// TIA Portal project "HEAT-1-CADIZ-V30" (V20) (continued)
VAR_GLOBAL   // PLC tag table "Robot Position"
   "tcpPosIniX_00" AT %I632.0 : Bool;   // $OUT[257]
   "tcpPosIniX_01" AT %I632.1 : Bool;
   "tcpPosIniX_02" AT %I632.2 : Bool;
   "tcpPosIniX_03" AT %I632.3 : Bool;
   "tcpPosIniX_04" AT %I632.4 : Bool;
   "tcpPosIniX_05" AT %I632.5 : Bool;
   "tcpPosIniX_06" AT %I632.6 : Bool;
   "tcpPosIniX_07" AT %I632.7 : Bool;
   "tcpPosIniX_08" AT %I633.0 : Bool;
   "tcpPosIniX_09" AT %I633.1 : Bool;
   "tcpPosIniX_10" AT %I633.2 : Bool;
   "tcpPosIniX_11" AT %I633.3 : Bool;
   "tcpPosIniX_12" AT %I633.4 : Bool;
   "tcpPosIniX_13" AT %I633.5 : Bool;
   "tcpPosIniX_14" AT %I633.6 : Bool;
   "tcpPosIniX_15" AT %I633.7 : Bool;
   "tcpPosIniX_16" AT %I634.0 : Bool;
   "tcpPosIniX_17" AT %I634.1 : Bool;
   "tcpPosIniX_18" AT %I634.2 : Bool;
   "tcpPosIniX_19" AT %I634.3 : Bool;
   "tcpPosIniX_20" AT %I634.4 : Bool;
   "tcpPosIniX_21" AT %I634.5 : Bool;
   "tcpPosIniX_22" AT %I634.6 : Bool;
   "tcpPosIniX_23" AT %I634.7 : Bool;
   "tcpPosIniX_24" AT %I635.0 : Bool;
   "tcpPosIniX_25" AT %I635.1 : Bool;
   "tcpPosIniX_26" AT %I635.2 : Bool;
   "tcpPosIniX_27" AT %I635.3 : Bool;
   "tcpPosIniX_28" AT %I635.4 : Bool;
   "tcpPosIniX_29" AT %I635.5 : Bool;
   "tcpPosIniX_30" AT %I635.6 : Bool;
   "tcpPosIniX_31" AT %I635.7 : Bool;
   "tcpPosIniY_00" AT %I636.0 : Bool;
   "tcpPosIniY_01" AT %I636.1 : Bool;
   "tcpPosIniY_02" AT %I636.2 : Bool;
   "tcpPosIniY_03" AT %I636.3 : Bool;
   "tcpPosIniY_04" AT %I636.4 : Bool;
   "tcpPosIniY_05" AT %I636.5 : Bool;
   "tcpPosIniY_06" AT %I636.6 : Bool;
   "tcpPosIniY_07" AT %I636.7 : Bool;
   "tcpPosIniY_08" AT %I637.0 : Bool;
   "tcpPosIniY_09" AT %I637.1 : Bool;
   "tcpPosIniY_10" AT %I637.2 : Bool;
   "tcpPosIniY_11" AT %I637.3 : Bool;
   "tcpPosIniY_12" AT %I637.4 : Bool;
   "tcpPosIniY_13" AT %I637.5 : Bool;
   "tcpPosIniY_14" AT %I637.6 : Bool;
   "tcpPosIniY_15" AT %I637.7 : Bool;
   "tcpPosIniY_16" AT %I638.0 : Bool;
   "tcpPosIniY_17" AT %I638.1 : Bool;
   "tcpPosIniY_18" AT %I638.2 : Bool;
   "tcpPosIniY_19" AT %I638.3 : Bool;
   "tcpPosIniY_20" AT %I638.4 : Bool;
   "tcpPosIniY_21" AT %I638.5 : Bool;
   "tcpPosIniY_22" AT %I638.6 : Bool;
   "tcpPosIniY_23" AT %I638.7 : Bool;
   "tcpPosIniY_24" AT %I639.0 : Bool;
   "tcpPosIniY_25" AT %I639.1 : Bool;
   "tcpPosIniY_26" AT %I639.2 : Bool;
   "tcpPosIniY_27" AT %I639.3 : Bool;
   "tcpPosIniY_28" AT %I639.4 : Bool;
   "tcpPosIniY_29" AT %I639.5 : Bool;
   "tcpPosIniY_30" AT %I639.6 : Bool;
   "tcpPosIniY_31" AT %I639.7 : Bool;
   "tcpPosIniZ_00" AT %I640.0 : Bool;
   "tcpPosIniZ_01" AT %I640.1 : Bool;
   "tcpPosIniZ_02" AT %I640.2 : Bool;
   "tcpPosIniZ_03" AT %I640.3 : Bool;
   "tcpPosIniZ_04" AT %I640.4 : Bool;
   "tcpPosIniZ_05" AT %I640.5 : Bool;
   "tcpPosIniZ_06" AT %I640.6 : Bool;
   "tcpPosIniZ_07" AT %I640.7 : Bool;
   "tcpPosIniZ_08" AT %I641.0 : Bool;
   "tcpPosIniZ_09" AT %I641.1 : Bool;
   "tcpPosIniZ_10" AT %I641.2 : Bool;
   "tcpPosIniZ_11" AT %I641.3 : Bool;
   "tcpPosIniZ_12" AT %I641.4 : Bool;
   "tcpPosIniZ_13" AT %I641.5 : Bool;
   "tcpPosIniZ_14" AT %I641.6 : Bool;
   "tcpPosIniZ_15" AT %I641.7 : Bool;
   "tcpPosIniZ_16" AT %I642.0 : Bool;
   "tcpPosIniZ_17" AT %I642.1 : Bool;
   "tcpPosIniZ_18" AT %I642.2 : Bool;
   "tcpPosIniZ_19" AT %I642.3 : Bool;
   "tcpPosIniZ_20" AT %I642.4 : Bool;
   "tcpPosIniZ_21" AT %I642.5 : Bool;
   "tcpPosIniZ_22" AT %I642.6 : Bool;
   "tcpPosIniZ_23" AT %I642.7 : Bool;
   "tcpPosIniZ_24" AT %I643.0 : Bool;
   "tcpPosIniZ_25" AT %I643.1 : Bool;
   "tcpPosIniZ_26" AT %I643.2 : Bool;
   "tcpPosIniZ_27" AT %I643.3 : Bool;
   "tcpPosIniZ_28" AT %I643.4 : Bool;
   "tcpPosIniZ_29" AT %I643.5 : Bool;
   "tcpPosIniZ_30" AT %I643.6 : Bool;
   "tcpPosIniZ_31" AT %I643.7 : Bool;
   "e1PosIni_00" AT %I644.0 : Bool;
   "e1PosIni_01" AT %I644.1 : Bool;
   "e1PosIni_02" AT %I644.2 : Bool;
   "e1PosIni_03" AT %I644.3 : Bool;
   "e1PosIni_04" AT %I644.4 : Bool;
   "e1PosIni_05" AT %I644.5 : Bool;
   "e1PosIni_06" AT %I644.6 : Bool;
   "e1PosIni_07" AT %I644.7 : Bool;
   "e1PosIni_08" AT %I645.0 : Bool;
   "e1PosIni_09" AT %I645.1 : Bool;
   "e1PosIni_10" AT %I645.2 : Bool;
   "e1PosIni_11" AT %I645.3 : Bool;
   "e1PosIni_12" AT %I645.4 : Bool;
   "e1PosIni_13" AT %I645.5 : Bool;
   "e1PosIni_14" AT %I645.6 : Bool;
   "e1PosIni_15" AT %I645.7 : Bool;
   "e1PosIni_16" AT %I646.0 : Bool;
   "e1PosIni_17" AT %I646.1 : Bool;
   "e1PosIni_18" AT %I646.2 : Bool;
   "e1PosIni_19" AT %I646.3 : Bool;
   "e1PosIni_20" AT %I646.4 : Bool;
   "e1PosIni_21" AT %I646.5 : Bool;
   "e1PosIni_22" AT %I646.6 : Bool;
   "e1PosIni_23" AT %I646.7 : Bool;
   "e1PosIni_24" AT %I647.0 : Bool;
   "e1PosIni_25" AT %I647.1 : Bool;
   "e1PosIni_26" AT %I647.2 : Bool;
   "e1PosIni_27" AT %I647.3 : Bool;
   "e1PosIni_28" AT %I647.4 : Bool;
   "e1PosIni_29" AT %I647.5 : Bool;
   "e1PosIni_30" AT %I647.6 : Bool;
   "e1PosIni_31" AT %I647.7 : Bool;
   "tcpPosFinX_00" AT %I648.0 : Bool;
   "tcpPosFinX_01" AT %I648.1 : Bool;
   "tcpPosFinX_02" AT %I648.2 : Bool;
   "tcpPosFinX_03" AT %I648.3 : Bool;
   "tcpPosFinX_04" AT %I648.4 : Bool;
   "tcpPosFinX_05" AT %I648.5 : Bool;
   "tcpPosFinX_06" AT %I648.6 : Bool;
   "tcpPosFinX_07" AT %I648.7 : Bool;
   "tcpPosFinX_08" AT %I649.0 : Bool;
   "tcpPosFinX_09" AT %I649.1 : Bool;
   "tcpPosFinX_10" AT %I649.2 : Bool;
   "tcpPosFinX_11" AT %I649.3 : Bool;
   "tcpPosFinX_12" AT %I649.4 : Bool;
   "tcpPosFinX_13" AT %I649.5 : Bool;
   "tcpPosFinX_14" AT %I649.6 : Bool;
   "tcpPosFinX_15" AT %I649.7 : Bool;
   "tcpPosFinX_16" AT %I650.0 : Bool;
   "tcpPosFinX_17" AT %I650.1 : Bool;
   "tcpPosFinX_18" AT %I650.2 : Bool;
   "tcpPosFinX_19" AT %I650.3 : Bool;
   "tcpPosFinX_20" AT %I650.4 : Bool;
   "tcpPosFinX_21" AT %I650.5 : Bool;
   "tcpPosFinX_22" AT %I650.6 : Bool;
   "tcpPosFinX_23" AT %I650.7 : Bool;
   "tcpPosFinX_24" AT %I651.0 : Bool;
   "tcpPosFinX_25" AT %I651.1 : Bool;
   "tcpPosFinX_26" AT %I651.2 : Bool;
   "tcpPosFinX_27" AT %I651.3 : Bool;
   "tcpPosFinX_28" AT %I651.4 : Bool;
   "tcpPosFinX_29" AT %I651.5 : Bool;
   "tcpPosFinX_30" AT %I651.6 : Bool;
   "tcpPosFinX_31" AT %I651.7 : Bool;
   "tcpPosFinY_00" AT %I652.0 : Bool;
   "tcpPosFinY_01" AT %I652.1 : Bool;
   "tcpPosFinY_02" AT %I652.2 : Bool;
   "tcpPosFinY_03" AT %I652.3 : Bool;
   "tcpPosFinY_04" AT %I652.4 : Bool;
   "tcpPosFinY_05" AT %I652.5 : Bool;
   "tcpPosFinY_06" AT %I652.6 : Bool;
   "tcpPosFinY_07" AT %I652.7 : Bool;
   "tcpPosFinY_08" AT %I653.0 : Bool;
   "tcpPosFinY_09" AT %I653.1 : Bool;
   "tcpPosFinY_10" AT %I653.2 : Bool;
   "tcpPosFinY_11" AT %I653.3 : Bool;
   "tcpPosFinY_12" AT %I653.4 : Bool;
   "tcpPosFinY_13" AT %I653.5 : Bool;
   "tcpPosFinY_14" AT %I653.6 : Bool;
   "tcpPosFinY_15" AT %I653.7 : Bool;
   "tcpPosFinY_16" AT %I654.0 : Bool;
   "tcpPosFinY_17" AT %I654.1 : Bool;
   "tcpPosFinY_18" AT %I654.2 : Bool;
   "tcpPosFinY_19" AT %I654.3 : Bool;
   "tcpPosFinY_20" AT %I654.4 : Bool;
   "tcpPosFinY_21" AT %I654.5 : Bool;
   "tcpPosFinY_22" AT %I654.6 : Bool;
   "tcpPosFinY_23" AT %I654.7 : Bool;
   "tcpPosFinY_24" AT %I655.0 : Bool;
   "tcpPosFinY_25" AT %I655.1 : Bool;
   "tcpPosFinY_26" AT %I655.2 : Bool;
   "tcpPosFinY_27" AT %I655.3 : Bool;
   "tcpPosFinY_28" AT %I655.4 : Bool;
   "tcpPosFinY_29" AT %I655.5 : Bool;
   "tcpPosFinY_30" AT %I655.6 : Bool;
   "tcpPosFinY_31" AT %I655.7 : Bool;
   "tcpPosE1_01" AT %I628.0 : Bool;
   "tcpPosE1_02" AT %I628.1 : Bool;
   "tcpPosE1_03" AT %I628.2 : Bool;
   "tcpPosE1_04" AT %I628.3 : Bool;
   "tcpPosE1_05" AT %I628.4 : Bool;
   "tcpPosE1_06" AT %I628.5 : Bool;
   "tcpPosE1_07" AT %I628.6 : Bool;
   "tcpPosE1_08" AT %I628.7 : Bool;
   "tcpPosE1_09" AT %I629.0 : Bool;
   "tcpPosE1_10" AT %I629.1 : Bool;
   "tcpPosE1_11" AT %I629.2 : Bool;
   "tcpPosE1_12" AT %I629.3 : Bool;
   "tcpPosE1_13" AT %I629.4 : Bool;
   "tcpPosE1_14" AT %I629.5 : Bool;
   "tcpPosE1_15" AT %I629.6 : Bool;
   "tcpPosE1_16" AT %I629.7 : Bool;
   "tcpPosE1_17" AT %I630.0 : Bool;
   "tcpPosE1_18" AT %I630.1 : Bool;
   "tcpPosE1_19" AT %I630.2 : Bool;
   "tcpPosE1_20" AT %I630.3 : Bool;
   "tcpPosE1_21" AT %I630.4 : Bool;
   "tcpPosE1_22" AT %I630.5 : Bool;
   "tcpPosE1_23" AT %I630.6 : Bool;
   "tcpPosE1_24" AT %I630.7 : Bool;
   "tcpPosE1_25" AT %I631.0 : Bool;
   "tcpPosE1_26" AT %I631.1 : Bool;
   "tcpPosE1_27" AT %I631.2 : Bool;
   "tcpPosE1_28" AT %I631.3 : Bool;
   "tcpPosE1_29" AT %I631.4 : Bool;
   "tcpPosE1_30" AT %I631.5 : Bool;
   "tcpPosE1_31" AT %I631.6 : Bool;
   "tcpPosE1_32" AT %I631.7 : Bool;
   "tcpPosIniX_rawLe32" AT %ID632 : DWord;
   "tcpPosIniY_rawLe32" AT %ID636 : DWord;
   "tcpPosIniZ_rawLe32" AT %ID640 : DWord;
   "tcpPosFinX_rawLe32" AT %ID648 : DWord;
   "tcpPosFinY_rawLe32" AT %ID652 : DWord;
   "e1_rawLe32" AT %ID628 : DWord;
   "e1PosIni_rawLe32" AT %ID644 : DWord;
   "tcpPosFinZ_rawLe32" AT %ID656 : DWord;
   "e1PosFin_rawLe32" AT %ID660 : DWord;
END_VAR

VAR_GLOBAL   // PLC tag table "Tool Change"
   "dockSensorToolYugoInPosition" AT %I150.0 : Bool;   // DETECTOR_YUGO_LP
   "dockSensorCoverYugoClosed" AT %I150.1 : Bool;   // TAPA_CERRADA_YUGO_LP
   "dockSensorCoverOpenYugo" AT %I160.0 : Bool;   // TAPA_ABIERTA_YUGO_LP
   "dockValveV2UnlockOnYugo" AT %Q171.2 : Bool;   // SOLTAR_HERRAMIENTA_YUGO_LP / CAMBIA A FALSE
   "dockValveCoverOpenOnYugo" AT %Q170.0 : Bool;   // ABRIR_TAPA_YUGO_LP
   "dockValveCoverCloseOnYugo" AT %Q170.1 : Bool;   // CERRAR_TAPA_YUGO_LP
   "robotSensorMpsUnlocked" AT %I200.0 : Bool;   // INTERCAMBIO_DESBLOQUEADO_LR
   "robotSensorMpsLocked" AT %I200.1 : Bool;   // INTERCAMBIO_BLOQUEADO_LR
   "robotSensorMpsCoupled" AT %I200.2 : Bool;   // HERRAMIENTA_PUESTA_LR /AL COLOCAR METAL
   "robotSensorMpsCtrlAirPressureOk" AT %I200.3 : Bool;   // PRESION_CORRECTA_LR
   "toolReqId_01" AT %Q618.1 : Bool;   // INKUKA_DETECTOR_HERRAMIENTA
   "toolReqId_02" AT %Q618.2 : Bool;   // INKUKA_TAPA_CERRADA_YUGO
   "toolReqId_03" AT %Q618.3 : Bool;   // INKUKA_TAPA_ABIERTA_YUGO
   "toolReqId_04" AT %Q618.4 : Bool;   // INKUKA_INTERCAMBIO_DESBLOQUEADO
   "toolReqId_05" AT %Q618.5 : Bool;   // INKUKA_INTERCAMBIO_BLOQUEADO
   "toolReqId_06" AT %Q618.6 : Bool;   // INKUKA_HERRAMIENTA_PUESTA /AL COLOCAR util met
   "toolReqId_07" AT %Q618.7 : Bool;
   "kukaCmdUnlockMpsYugo" AT %I696.0 : Bool;   // OUTKUKA_SOLTAR_HERRAMIENTA_YUGO
   "kukaCmdOpenCover" AT %I696.1 : Bool;   // OUTKUKA_ABRIR_TAPA_YUGO
   "kukaCmdCloseCover" AT %I696.2 : Bool;   // OUTKUKA_CERRAR_TAPA_YUGO
   "V1_B14_S2" AT %Q0.0 : Bool;   // Anticolision - OPR
   "V1_B12_S4" AT %Q0.1 : Bool;   // Mps Bloqueo SIL 2
   "V2_B14_S2" AT %Q0.2 : Bool;
   "V2_B12_S4" AT %Q0.3 : Bool;
   "toolReqId_00" AT %Q618.0 : Bool;
   "toolReqId_08" AT %Q619.0 : Bool;
   "toolReqId_09" AT %Q619.1 : Bool;
   "toolReqId_10" AT %Q619.2 : Bool;
   "toolReqId_11" AT %Q619.3 : Bool;
   "toolReqId_12" AT %Q619.4 : Bool;
   "toolReqId_13" AT %Q619.5 : Bool;
   "toolReqId_14" AT %Q619.6 : Bool;
   "toolReqId_15" AT %Q619.7 : Bool;
   "toolReqId" AT %QW618 : Word;
   "baseReqId" AT %QW620 : Word;
   "kukaFeedbackDockToolYugoInPosition" AT %Q696.4 : Bool;   // $IN[773]
   "kukaFeedbackDockYugoCoverClosed" AT %Q696.5 : Bool;
   "kukaFeedbackDockYugoCoverOpen" AT %Q696.6 : Bool;
   "kukaFeedbackRobotMpsUnlocked" AT %Q696.0 : Bool;   // $IN[769]
   "kukaFeedbackRobotMpsLocked" AT %Q696.1 : Bool;
   "kukaFeedbackRobotMpsCoupled" AT %Q696.2 : Bool;
   "kukaFeedbackRobotMpsCtrlAirPressureOk" AT %Q696.3 : Bool;
   "dockValveV2UnlockOnPepa" AT %Q171.4 : Bool;   // SOLTAR_HERRAMIENTA_PEPA
   "dockSensorToolPepaInPosition" AT %I150.2 : Bool;
   "kukaCmdSafeForChange" AT %I696.3 : Bool;   // $OUT[772]
   "kukaCmdUnlockMpsPepa" AT %I696.4 : Bool;   // $OUT[773]
   "kukaCmdOpenCoverPepa" AT %I696.5 : Bool;   // $OUT[774]
   "kukaCmdUnlockMpsMarker" AT %I696.7 : Bool;   // $OUT[775]
   "kukaCmdOpenCoverMarker" AT %I697.0 : Bool;   // $OUT[776]
   "kukaCmdCloseCoverMarker" AT %I697.1 : Bool;   // $OUT[777]
   "kukaCmdUnlockMpsGocator" AT %I697.2 : Bool;
   "kukaCmdOpenCoverGocator" AT %I697.3 : Bool;
   "kukaCmdCloseCoverGocator" AT %I697.4 : Bool;
   "kukaCmdCloseCoverPepa" AT %I696.6 : Bool;
   "kukaCmdUnlockMpsPole" AT %I697.5 : Bool;
   "kukaCmdOpenCoverPole" AT %I697.6 : Bool;
   "kukaCmdCloseCoverPole" AT %I697.7 : Bool;
   "kukaFeedbackDockToolPepaInPosition" AT %Q696.7 : Bool;
   "kukaFeedbackDockPepaCoverClosed" AT %Q697.0 : Bool;
   "kukaFeedbackDockPepaCoverOpen" AT %Q697.1 : Bool;
   "kukaFeedbackDockToolMarkerInPosition" AT %Q697.2 : Bool;
   "kukaFeedbackDockMarkerCoverClosed" AT %Q697.3 : Bool;
   "kukaFeedbackDockMarkerCoverOpen" AT %Q697.4 : Bool;
   "kukaFeedbackDockToolGocatorInPosition" AT %Q697.5 : Bool;
   "kukaFeedbackDockGocatorCoverClosed" AT %Q697.6 : Bool;
   "kukaFeedbackDockGocatorCoverOpen" AT %Q697.7 : Bool;
   "kukaFeedbackDockToolPoleInPosition" AT %Q698.0 : Bool;
   "kukaFeedbackDockPoleCoverClosed" AT %Q698.1 : Bool;
   "kukaFeedbackDockPoleCoverOpen" AT %Q698.2 : Bool;
   "dockSensorCoverPepaClosed" AT %I150.3 : Bool;
   "dockSensorToolPoleInPosition" AT %I150.4 : Bool;
   "dockSensorToolMarkerInPosition" AT %I150.6 : Bool;
   "dockSensorToolGocatorInPosition" AT %I151.0 : Bool;
   "pruebaHerramienta2enStand" AT %I151.2 : Bool;
   "dockSensorCoverGocatorClosed" AT %I151.1 : Bool;
   "pruebaHerramienta3enStand" AT %I151.3 : Bool;
   "pruebaHerramienta4enStand" AT %I151.4 : Bool;
   "dockSensorCoverMarkerClosed" AT %I150.7 : Bool;
   "dockSensorCoverPOLEClosed" AT %I150.5 : Bool;
   "toolIdProxy1" AT %I201.0 : Bool;
   "toolIdProxy2" AT %I201.1 : Bool;
   "toolIdProxy3" AT %I201.2 : Bool;
   "toolIdProxy4" AT %I201.3 : Bool;
   "dockSensorCoverOpenPepa" AT %I160.1 : Bool;
   "dockSensorCoverOpenPOLE" AT %I160.2 : Bool;
   "dockSensorCoverOpenMarker" AT %I160.3 : Bool;
   "dockSensorCoverOpenGocator" AT %I160.4 : Bool;
   "dockValveV2UnlockOnMarker" AT %Q180.0 : Bool;
   "dockValveV2UnlockOnGocator" AT %Q180.2 : Bool;
END_VAR

VAR_GLOBAL   // PLC tag table "General"
   "ALM_PRESS_SENSOR" AT %I10.0 : Bool;   // Pressure-sensor alarm
END_VAR

VAR_GLOBAL   // PLC tag table "CUBA"
   "Sensor_plato_giro_1" AT %I410.0 : Bool;
   "Sensor_Plato_giro_2" AT %I410.1 : Bool;
   "Sensor_plato_giro_3" AT %I410.2 : Bool;
   "--" AT %I410.3 : Bool;
   "SENSOR_DSBG_BASTIDOR_ABAJO_1" AT %I410.4 : Bool;
   "SENSOR_DSBG_BASTIDOR_ARRIBA_1" AT %I410.5 : Bool;
   "SENSOR_DSBG_BASTIDOR_ABAJO_2" AT %I410.6 : Bool;
   "SENSOR_DSBG_BASTIDOR_ARRIBA_2" AT %I410.7 : Bool;
   "Sensor_ADN_bastidor_bloqueado_1" AT %I411.0 : Bool;
   "Sensor_ADN_bastidor_bdesloqueado_1" AT %I411.1 : Bool;
   "Sensor_ADN_bastidor_bloqueado_2" AT %I411.2 : Bool;
   "Sensor_ADN_bastidor_desbloqueado_2" AT %I411.3 : Bool;
   "SENSOR_CENTRO_CUBA_ABAJO_1" AT %I411.4 : Bool;
   "SENSOR_CENTRO_CUBA_ARRIBA_1" AT %I411.5 : Bool;
   "SENSOR_CENTRO_CUBA_ABAJO_2" AT %I411.6 : Bool;
   "PULSADOR_SUBIR_1" AT %I412.0 : Bool;
   "PULSADOR_BAJAR_1" AT %I412.1 : Bool;
   "PULSADOR_SUBIR_2" AT %I412.2 : Bool;
   "PULSADOR_BAJAR_2" AT %I412.3 : Bool;
   "VALVULA_52_BIESTABLE_11" AT %Q420.0 : Bool;
   "VALVULA_52_BIESTABLE_12" AT %Q420.1 : Bool;
   "VALVULA_52_BIESTABLE_21" AT %Q420.2 : Bool;
   "VALVULA_52_BIESTABLE_22" AT %Q420.3 : Bool;
   "VÁLVULA_52_MONOESTABLE_1" AT %Q420.4 : Bool;
   "VÁLVULA_52_MONOESTABLE_2" AT %Q420.5 : Bool;
   "VÁLVULA_52_MONOESTABLE_3" AT %Q420.6 : Bool;
   "VÁLVULA_52_MONOESTABLE_4" AT %Q420.7 : Bool;
   "VÁLVULA_52_MONOESTABLE_5" AT %Q421.0 : Bool;
   "SENSOR_CENTRO_CUBA_ARRIBA_2" AT %I411.7 : Bool;
   "Libre" AT %I412.4 : Bool;
   "Libre(1)" AT %I412.5 : Bool;
   "libre(2)" AT %I412.6 : Bool;
   "libre(3)" AT %I412.7 : Bool;
   "Sensor_nivel_cuba_superior" AT %I413.0 : Bool;
   "Sensor_nivel_cuba_superior(1)" AT %I413.1 : Bool;
   "Sensor_nivel_cuba_medio(2)" AT %I413.2 : Bool;
   "Sensor_nivel_cuba_medio(1)" AT %I413.3 : Bool;
   "Sensor_nivel_cuba_inferior(1)" AT %I413.4 : Bool;
   "Sensor_nivel_cuba_inferior(2)" AT %I413.5 : Bool;
   "libre(4)" AT %I413.6 : Bool;
   "libre(5)" AT %I413.7 : Bool;
   "VÁLVULA_52_MONOESTABLE_6" AT %Q421.1 : Bool;
   "VÁLVULA_52_MONOESTABLE_7" AT %Q421.2 : Bool;
   "VÁLVULA_52_MONOESTABLE_8" AT %Q421.3 : Bool;
   "VÁLVULA_52_MONOESTABLE_9" AT %Q421.4 : Bool;
   "VÁLVULA_52_MONOESTABLE_10" AT %Q421.5 : Bool;
   "VÁLVULA_52_MONOESTABLE_11" AT %Q421.6 : Bool;
   "VÁLVULA_52_MONOESTABLE_12" AT %Q421.7 : Bool;
   "VÁLVULA_52_MONOESTABLE_13" AT %Q422.0 : Bool;
   "VÁLVULA_52_MONOESTABLE_14" AT %Q422.1 : Bool;
   "VÁLVULA_52_MONOESTABLE_15" AT %Q422.2 : Bool;
   "VÁLVULA_52_MONOESTABLE_16" AT %Q422.3 : Bool;
   "VÁLVULA_52_MONOESTABLE_17" AT %Q422.4 : Bool;
   "VÁLVULA_52_MONOESTABLE_18" AT %Q422.5 : Bool;
   "VÁLVULA_52_MONOESTABLE_19" AT %Q422.6 : Bool;
   "VÁLVULA_52_MONOESTABLE_20" AT %Q422.7 : Bool;
   "VÁLVULA_52_MONOESTABLE_21" AT %Q423.0 : Bool;
   "VÁLVULA_52_MONOESTABLE_22" AT %Q423.1 : Bool;
   "VÁLVULA_52_MONOESTABLE_23" AT %Q423.2 : Bool;
   "VÁLVULA_52_MONOESTABLE_24" AT %Q423.3 : Bool;
   "VÁLVULA_52_MONOESTABLE_25" AT %Q423.4 : Bool;
   "VÁLVULA_52_MONOESTABLE_26" AT %Q423.5 : Bool;
   "VÁLVULA_52_MONOESTABLE_27" AT %Q423.6 : Bool;
   "VÁLVULA_52_MONOESTABLE_28" AT %Q423.7 : Bool;
   "CMD_TANK_DRAIN" AT %Q30.1 : Bool;   // VACIAR CUBA
   "CMD_TANK_FILL" AT %Q30.0 : Bool;   // LLENAR CUBA
   "RECIRCULACION" AT %Q30.2 : Bool;   // CONMUTADOR MANUAL / cambiado a recirculacion
   "MODE_WATER_AUTO" AT %Q30.3 : Bool;   // CONMUTADOR AUTO_NO_ESTA
   "ACTIVAR_ELECTROIMAN" AT %Q30.4 : Bool;   // ACTIVAR ELECTRO_IMAN_PUERTA
END_VAR

VAR_GLOBAL   // PLC tag table "ROBOT_SAFE_OPERATION"
   "NHL" AT %I500.0 : Bool;   // Parada de eergencia local
   "AF" AT %I500.1 : Bool;   // habilitacion de accionamientos
   "FF" AT %I500.2 : Bool;   // liberacion de movimiento
   "ZS" AT %I500.3 : Bool;   // validacion ext
   "PE" AT %I500.4 : Bool;   // conectar la periferia
   "AUT" AT %I500.5 : Bool;   // modo servicio automatico-ext
   "T1" AT %I500.6 : Bool;   // modo servicio t1
   "T2" AT %I500.7 : Bool;   // modo servicio t2
   "NHE" AT %I501.0 : Bool;   // parada emergencia externa
   "BSQ" AT %I501.1 : Bool;   // proteccion contra operario confirmada
   "SHS1" AT %I501.2 : Bool;   // parada de seguridad 1
   "SHS2" AT %I501.3 : Bool;   // parada de seguridad 2
   "RESERVADO_1" AT %I501.4 : Bool;
   "RESERVADO_2" AT %I501.5 : Bool;
   "PSA" AT %I501.6 : Bool;   // interfaz de seguridad activa
   "SP" AT %I501.7 : Bool;   // sistema powerdown
   "SO" AT %I502.0 : Bool;   // supervisiones seguras activas
   "RR" AT %I502.1 : Bool;   // referencia robot
   "JF" AT %I502.2 : Bool;   // error de ajuste
   "VRED" AT %I502.3 : Bool;   // velocidad reducida
   "SBHS1" AT %I502.4 : Bool;   // parada de servicio segura grupo de ejes 1
   "SBHS2" AT %I502.5 : Bool;   // parada de servicio segura grupo de ejes 2
   "SBHS3" AT %I502.6 : Bool;   // parada de servicio segura grupo de ejes 3
   "SBHS4" AT %I502.7 : Bool;   // parada de servicio segura grupo de ejes 4
   "SBHS5" AT %I503.0 : Bool;   // parada de servicio segura grupo de ejes 5
   "SBHS6" AT %I503.1 : Bool;   // parada de servicio segura grupo de ejes 6
   "SOS" AT %I503.2 : Bool;   // parada safe operation
   "RESERVADO_3" AT %I503.3 : Bool;
   "RESERVADO_4" AT %I503.4 : Bool;
   "RESERVADO_5" AT %I503.5 : Bool;
   "RESERVADO_6" AT %I503.6 : Bool;
   "RESERVADO_7" AT %I503.7 : Bool;
   "MR1" AT %I504.0 : Bool;   // espacio de aviso 1
   "MR2" AT %I504.1 : Bool;   // espacio de aviso 2
   "MR3" AT %I504.2 : Bool;   // espacio de aviso 3
   "MR4" AT %I504.3 : Bool;   // espacio de aviso 4
   "MR5" AT %I504.4 : Bool;   // espacio de aviso 5
   "MR6" AT %I504.5 : Bool;   // espacio de aviso 6
   "MR7" AT %I504.6 : Bool;   // espacio de aviso 7
   "MR8" AT %I504.7 : Bool;   // espacio de aviso 8
   "MR9" AT %I505.0 : Bool;   // espacio de aviso 9
   "MR10" AT %I505.1 : Bool;   // espacio de aviso 10
   "MR11" AT %I505.2 : Bool;   // espacio de aviso 11
   "MR12" AT %I505.3 : Bool;   // espacio de aviso 12
   "MR13" AT %I505.4 : Bool;   // espacio de aviso 13
   "MR14" AT %I505.5 : Bool;   // espacio de aviso 14
   "MR15" AT %I505.6 : Bool;   // espacio de aviso 15
   "MR16" AT %I505.7 : Bool;   // espacio de aviso 16
   "RESERVADO_8" AT %I506.0 : Bool;
   "RESERVADO_9" AT %I506.1 : Bool;
   "RESERVADO_10" AT %I506.2 : Bool;
   "RESERVADO_11" AT %I506.3 : Bool;
   "RESERVADO_12" AT %I506.4 : Bool;
   "RESERVADO_13" AT %I506.5 : Bool;
   "RESERVADO_14" AT %I506.6 : Bool;
   "RESERVADO_15" AT %I506.7 : Bool;
   "RESERVADO_16" AT %I507.0 : Bool;
   "RESERVADO_17" AT %I507.1 : Bool;
   "RESERVADO_18" AT %I507.2 : Bool;
   "RESERVADO_19" AT %I507.3 : Bool;
   "RESERVADO_20" AT %I507.4 : Bool;
   "RESERVADO_21" AT %I507.5 : Bool;
   "RESERVADO_22" AT %I507.6 : Bool;
   "RESERVADO_23" AT %I507.7 : Bool;
   "RES1 (reservado)" AT %Q500.0 : Bool;
   "NHE – E‑Stop externo" AT %Q500.1 : Bool;   // E‑Stop externo
   "BS – Puerta cerrada" AT %Q500.2 : Bool;   // Puerta cerrada
   "QBS – Ack puerta" AT %Q500.3 : Bool;   // confirmacion de puerta cerrada
   "SHS1 – Stop 1" AT %Q500.4 : Bool;   // parada de seguridad 1
   "SHS2 – Stop 2" AT %Q500.5 : Bool;   // parada de seguridad 2
   "RES6" AT %Q500.6 : Bool;
   "RES7" AT %Q500.7 : Bool;
   "US2 – 24 V US2" AT %Q501.0 : Bool;   // contactor de periferia
   "SBH" AT %Q501.1 : Bool;   // parada de servicio segura
   "RES11" AT %Q501.2 : Bool;
   "RES12" AT %Q501.3 : Bool;
   "RES13" AT %Q501.4 : Bool;
   "RES14" AT %Q501.5 : Bool;
   "RES15" AT %Q501.6 : Bool;
   "SPA – Power‑down Ack" AT %Q501.7 : Bool;   // Confirmacion de parada del controlador
   "JR" AT %Q502.0 : Bool;   // interruptor de referencia de ajuste
   "VRED_OUT" AT %Q502.1 : Bool;   // velocidad reducida
   "SBH_OUT_1" AT %Q502.2 : Bool;   // parada de servicio segura de grupo de ejes 1
   "SBH_OUT_2" AT %Q502.3 : Bool;   // parada de servicio segura de grupo de ejes 2
   "SBH_OUT_3" AT %Q502.4 : Bool;   // parada de servicio segura de grupo de ejes 3
   "SBH_OUT_4" AT %Q502.5 : Bool;   // parada de servicio segura de grupo de ejes 4
   "SBH_OUT_5" AT %Q502.6 : Bool;   // parada de servicio segura de grupo de ejes 5
   "SBH_OUT_6" AT %Q502.7 : Bool;   // parada de servicio segura de grupo de ejes 6
   "RES16" AT %Q503.0 : Bool;
   "RES17" AT %Q503.1 : Bool;
   "RES18" AT %Q503.2 : Bool;
   "RES19" AT %Q503.3 : Bool;
   "RES20" AT %Q503.4 : Bool;
   "RES21" AT %Q503.5 : Bool;
   "RES22" AT %Q503.6 : Bool;
   "RES23" AT %Q503.7 : Bool;
   "UER1" AT %Q504.0 : Bool;   // Zona de control1
   "UER2" AT %Q504.1 : Bool;   // Zona de control2
   "UER3" AT %Q504.2 : Bool;   // Zona de control3
   "UER4" AT %Q504.3 : Bool;   // Zona de control4
   "UER5" AT %Q504.4 : Bool;   // Zona de control5
   "UER6" AT %Q504.5 : Bool;   // Zona de control6
   "UER7" AT %Q504.6 : Bool;   // Zona de control7
   "UER8" AT %Q504.7 : Bool;   // Zona de control8
   "UER9" AT %Q505.0 : Bool;   // Zona de control9
   "UER10" AT %Q505.1 : Bool;   // Zona de control10
   "UER11" AT %Q505.2 : Bool;   // Zona de control11
   "UER12" AT %Q505.3 : Bool;   // Zona de control12
   "UER13" AT %Q505.4 : Bool;   // Zona de control13
   "UER14" AT %Q505.5 : Bool;   // Zona de control14
   "UER15" AT %Q505.6 : Bool;   // Zona de control15
   "UER16" AT %Q505.7 : Bool;   // Zona de control16
   "WZ1" AT %Q506.0 : Bool;   // Herramienta 1
   "WZ2" AT %Q506.1 : Bool;   // Herramienta 2
   "WZ3" AT %Q506.2 : Bool;   // Herramienta 3
   "WZ4" AT %Q506.3 : Bool;   // Herramienta 4
   "WZ5" AT %Q506.4 : Bool;   // Herramienta 5
   "WZ6" AT %Q506.5 : Bool;   // Herramienta 6
   "WZ7" AT %Q506.6 : Bool;   // Herramienta 7
   "WZ8" AT %Q506.7 : Bool;   // Herramienta 8
   "WZ9" AT %Q507.0 : Bool;   // Herramienta 9
   "WZ10" AT %Q507.1 : Bool;   // Herramienta 10
   "WZ11" AT %Q507.2 : Bool;   // Herramienta 11
   "WZ12" AT %Q507.3 : Bool;   // Herramienta 12
   "WZ13" AT %Q507.4 : Bool;   // Herramienta 13
   "WZ14" AT %Q507.5 : Bool;   // Herramienta 14
   "WZ15" AT %Q507.6 : Bool;   // Herramienta 15
   "WZ16" AT %Q507.7 : Bool;   // Herramienta 16
END_VAR

VAR_GLOBAL   // PLC tag table "SAFETY"
   "eStopButtonCabinet" AT %I40.0 : Bool;   // Emergency-Stop cabinet — 1oo2 result
   "eStopButtonTank" AT %I40.1 : Bool;   // Emergency-Stop tank — 1oo2 result
   "eStopButtonTankPartnerCh" AT %I41.1 : Bool;   // partner channel 1oo2 — do not use
   "eStopButtonWaterSystem" AT %I40.2 : Bool;   // Emergency-Stop water system — 1oo2 result
   "eStopButtonWaterSystemPartnerCh" AT %I41.2 : Bool;   // partner channel 1oo2 — do not use
   "eStopButtonHmiPanel" AT %I40.3 : Bool;   // Emergency-Stop HMI panel — 1oo2 result
   "eStopButtonHmiPanelPartnerCh" AT %I41.3 : Bool;   // partner channel 1oo2 — do not use
   "eStopButtonLightCurtain1" AT %I40.4 : Bool;   // Emergency-Stop light curtain 1 — 1oo2 resul
   "eStopButtonLightCurtain1PartnerCh" AT %I41.4 : Bool;   // partner channel 1oo2 — do not use
   "eStopButtonDoorPartnerCh" AT %I41.5 : Bool;   // partner channel 1oo2 — do not use
   "lightCurtain1Ossd1" AT %I50.0 : Bool;   // Z2 – LC 1 OSSD 1 (receiver)
   "lightCurtain1Ossd2" AT %I51.0 : Bool;   // Z2 – LC 1 OSSD 2 (receiver)
   "lightCurtain3Ossd1" AT %I50.1 : Bool;   // Z2 – LC 3 OSSD 1 (receiver)
   "lightCurtain3Ossd2" AT %I51.1 : Bool;   // Z2 – LC 3 OSSD 2 (receiver)
   "lightCurtain6Ossd1" AT %I50.2 : Bool;   // Z2 – LC 6 OSSD 1 (receiver)
   "lightCurtain6Ossd2" AT %I51.2 : Bool;   // Z2 – LC 6 OSSD 2 (receiver)
   "enableAccessReqSelector" AT %I50.3 : Bool;   // Rotary selector – enabless request access
   "DoorClosedCh1" AT %I50.6 : Bool;   // Safety door closed interlock – contact 1
   "resetDoorButton" AT %I50.7 : Bool;   // Reset push‑button
   "SAF_DOOR_CLSD_CH2" AT %I51.6 : Bool;   // Safety door closed interlock – contact 2
   "SAF_DOOR_UNLOCK_CH1" AT %Q60.0 : Bool;   // Unlock safety door – redundant output 1
   "SAF_GATE_UNLOCK_CH2" AT %Q60.2 : Bool;   // Unlock safety door – redundant output 2
   "accessReqButtonZone2" AT %I51.4 : Bool;   // Illuminated push-button – access request for zone 2
   "accessReqButtonZone3" AT %I51.5 : Bool;   // Illuminated push-button – access request for zone 3
   "accessReqButtonZone1" AT %I51.3 : Bool;   // Illuminated push-button – access request for zone 1
   "eStopButtonIslandRight1" AT %I300.1 : Bool;
   "buttonResetHmi" AT %I51.7 : Bool;
   "eStopButtonCabinetPartnerCh" AT %I41.0 : Bool;   // partner channel 1oo2 — do not use
   "PRESSURE_VALVE" AT %Q60.1 : Bool;
   "Door_output_1" AT %I50.4 : Bool;
   "Door_Output_2" AT %I50.5 : Bool;
   "eStopButtonDoor" AT %I40.5 : Bool;   // Emergency-Stop Door — 1oo2 result
END_VAR

TYPE "UDT_Dock"
   STRUCT
      Sensor : Struct
         CoverOpen : Bool;
         CoverClosed : Bool;
         ToolInPosition : Bool;
      END_STRUCT;
      Valve : Struct
         CoverOpenOn : Bool;
         CoverCloseOn : Bool;
         V2UnlockOn : Bool;
      END_STRUCT;
   END_STRUCT;
END_TYPE

TYPE "UDT_RobotMps"
   STRUCT
      Sensor : Struct
         Coupled : Bool;
         Locked : Bool;
         Unlocked : Bool;
         CtrlAirPressureOk : Bool;
      END_STRUCT;
   END_STRUCT;
END_TYPE

// folder: 10. System

DATA_BLOCK "HMI_CUBA_DB"   // DB17
{ S7_Optimized_Access := 'TRUE' }
VERSION : 0.1
// stored: InstanceOfName HMI_CUBA
"HMI_CUBA"
BEGIN
END_DATA_BLOCK

DATA_BLOCK "instKukaControlSeq_DB"   // DB20
{ S7_Optimized_Access := 'TRUE' }
VERSION : 0.1
// stored: InstanceOfName KukaControlSeq
"KukaControlSeq"
BEGIN
END_DATA_BLOCK

DATA_BLOCK "GIRO_POSITIVO_DB"   // DB27
{ S7_Optimized_Access := 'TRUE' }
VERSION : 0.1
// stored: InstanceOfName GIRO_POSITIVO
"GIRO_POSITIVO"
BEGIN
END_DATA_BLOCK

DATA_BLOCK "GIRO_NEGATIVO_1_DB"   // DB28
{ S7_Optimized_Access := 'TRUE' }
VERSION : 0.1
// stored: InstanceOfName GIRO_NEGATIVO_1
"GIRO_NEGATIVO_1"
BEGIN
END_DATA_BLOCK

// folder: 10. System/DbsInstancia

DATA_BLOCK "InstKukaControlSeq"   // DB14
{ S7_Optimized_Access := 'TRUE' }
VERSION : 0.1
// stored: InstanceOfName KukaControlSeq
"KukaControlSeq"
BEGIN
END_DATA_BLOCK

DATA_BLOCK "InstSupervisorSeq"   // DB15
{ S7_Optimized_Access := 'TRUE' }
VERSION : 0.1
// stored: InstanceOfName SupervisorSeq
"SupervisorSeq"
BEGIN
END_DATA_BLOCK

DATA_BLOCK "InstSeqManager"   // DB16
{ S7_Optimized_Access := 'TRUE' }
VERSION : 0.1
// stored: InstanceOfName SeqManager
"SeqManager"
BEGIN
END_DATA_BLOCK

DATA_BLOCK "AutoExtSeq_DB"   // DB18
{ S7_Optimized_Access := 'TRUE' }
VERSION : 0.1
// stored: InstanceOfName AutoExtSeq
"AutoExtSeq"
BEGIN
END_DATA_BLOCK

DATA_BLOCK "instSupervisorSeq_DB"   // DB21
{ S7_Optimized_Access := 'TRUE' }
VERSION : 0.1
// stored: InstanceOfName SupervisorSeq
"SupervisorSeq"
BEGIN
END_DATA_BLOCK

// folder: 10. System/DbsOpcUa

DATA_BLOCK "PlcStatus"   // DB4
{ S7_Optimized_Access := 'TRUE' }
VERSION : 0.1
   VAR
      "- FOR  KUKACONTROL-" : Bool;
      mode : Struct
         effective : UInt;
         ready : Bool;
      END_STRUCT;
      active : Struct
         baseId : UInt;
         toolId : UInt;
         profileId : UInt;
      END_STRUCT;
      exec : Struct
         ackSeq : UInt;
         accepted : Bool;
         busy : Bool;
         done : Bool;
         error : Bool;
         errorCode : UDInt;
         cancelAck : Bool;
         pauseAck : Bool;
         resumeAck : Bool;
         paused : Bool;
      END_STRUCT;
      pose : Struct
         tcpPosX_mm : LReal;
         tcpPosY_mm : LReal;
         tcpPosZ_mm : LReal;
         tcpOriA_deg : LReal;
         tcpOriB_deg : LReal;
         tcpOriC_deg : LReal;
         e1Pos_mm : LReal;
      END_STRUCT;
      teach : Struct
         startX_mm : LReal;
         startY_mm : LReal;
         startZ_mm : LReal;
         startE1_mm : LReal;
         startOk : Bool;
         endX_mm : LReal;
         endY_mm : LReal;
         endZ_mm : LReal;
         endE1_mm : LReal;
         endOk : Bool;
      END_STRUCT;
      systemArmed : Bool;
      robotInHome : Bool;
      robotInAutExt : Bool;
      heartbeatPlc : Bool;
      stepPlc : Int;
      plcOk : Bool := true;
      safetyOk : Bool := true;
      airOk : Bool := true;
      inspWaterOk : Bool := true;
      tankWaterOk : Bool := true;
      robotOk : Bool := true;
      acknowledge : Bool;
      carriageId : String;
      newCarriageId : Bool;
      idRunning : Bool;
      idOk : Bool;
      startUsReady : Bool;
      stopUsReady : Bool;
      paCheckReady : Bool;
      gainReady : Bool;
      tcgReady : Bool;
      idScan : String;
      pointOriginX : LReal;
      pointOriginY : LReal;
      pointOriginZ : LReal;
      xSize : LReal;
      ySize : LReal;
      scanRefStart : Bool;
      scanInspStart : Bool;
      markRunning : Bool;
      markState : Bool;
      breakUs : Bool;
      unbreakUs : Bool;
      robotRescanning : Bool;
      acknowledgeError : Bool;
   END_VAR
BEGIN
END_DATA_BLOCK

DATA_BLOCK "KukaControlCmd"   // DB5
{ S7_Optimized_Access := 'TRUE' }
VERSION : 0.1
   VAR
      code : UInt;
      seq : UInt;
      tcpTargetX_mm : LReal;
      tcpTargetY_mm : LReal;
      tcpTargetZ_mm : LReal;
      e1Target : LReal;
      toolRequestId : UInt;
      baseRequestId : UInt;
      profileRequestId : UInt;
      vel_mms : UInt;
      index_mm : UInt;
      apo_mm : LReal;
      programRequestId : UInt;
      cancelGo : Bool;
      pauseGo : Bool;
      resumeGo : Bool;
      mode : Struct
         request : UInt;
         reqSeq : UInt;
      END_STRUCT;
      scanPuntoInicialX : LReal;
      scanPuntoInicialY : LReal;
      scanPuntoInicialZ : LReal;
      scanPuntoInicialE1 : LReal;
      scanPuntoFinalX : LReal;
      scanPuntoFinalY : LReal;
      scanPuntoFinalZ : LReal;
      scanPuntoFinalE1 : LReal;
      carriageId : String;
      qrReady : Bool;
      drivesOn : Bool;
      extStart : Bool;
      confMess : Bool;
   END_VAR
BEGIN
END_DATA_BLOCK

DATA_BLOCK "SupervisorCmd"   // DB6
{ S7_Optimized_Access := 'TRUE' }
VERSION : 0.1
   VAR
      heartbeatSupervisor : Bool;
      stepSupervisor : Int;
      supervisorOk : Bool := true;
      stateUs : Bool;
      reqCarriageId : Bool;
      reqId : Bool;
      pns : Array[0..15] of String;
      referencePart : String;
      endEffector : Int;
      utTech : UInt;
      teachReq : Bool;
      paCheckReq : Bool;
      tcgReq : Bool;
      startUsRunning : Bool;
      stopUsRunning : Bool;
      elemState : Bool;
      elemRunning : Bool;
      balState : Bool;
      balRunning : Bool;
      gainState : Bool;
      gainRunning : Bool;
      tcgInProgress : Bool;
      tcgNextStep : Bool;
      tcgState : Bool;
      reqRefPart : Bool;
      reqStopCycle : Bool;
      reqTcgAdj : Bool;
      scanRefState : Bool;
      scanRefRunning : Bool;
      reqPreEval : Bool;
      reqIdentificationState : Bool;
      scanInspState : Bool;
      scanInsprunning : Bool;
      reqMark : Bool;
      reqVerif : Bool;
      pointCoordinates : LReal;
      goBack : Bool;
      rescanning : Bool;
      errorMessage : String;
      errorOcurred : Bool;
      gainAdjustmentReq : Bool;
   END_VAR
BEGIN
   pns[0] := 'M551B2810006-A01';
END_DATA_BLOCK

// folder: 10. System/Utilities

DATA_BLOCK "Utilidades"   // DB37
{ S7_Optimized_Access := 'TRUE' }
VERSION : 0.1
   VAR
      numProg : USInt;
   END_VAR
BEGIN
END_DATA_BLOCK

// folder: 20. Robot Services/AutoExt

DATA_BLOCK "instAutoExtSeq"   // DB7
{ S7_Optimized_Access := 'TRUE' }
VERSION : 0.1
// stored: InstanceOfName AutoExtSeq
"AutoExtSeq"
BEGIN
END_DATA_BLOCK

// folder: 20. Robot Services/DbsInstancia

DATA_BLOCK "InstTcpJogging"   // DB2
{ S7_Optimized_Access := 'TRUE' }
VERSION : 0.1
// stored: InstanceOfName TcpJogging
"TcpJogging"
BEGIN
END_DATA_BLOCK

DATA_BLOCK "ToolChangeFork_DB"   // DB8
{ S7_Optimized_Access := 'TRUE' }
VERSION : 0.1
// stored: InstanceOfName ToolChange
"ToolChange"
BEGIN
END_DATA_BLOCK

DATA_BLOCK "TcpPoseDecoderLe32_DB"   // DB10
{ S7_Optimized_Access := 'TRUE' }
VERSION : 0.1
// stored: InstanceOfName TcpPoseDecoderLe32
"TcpPoseDecoderLe32"
BEGIN
END_DATA_BLOCK

DATA_BLOCK "InstTcpTarget"   // DB13
{ S7_Optimized_Access := 'TRUE' }
VERSION : 0.1
// stored: InstanceOfName TcpTarget
"TcpTarget"
BEGIN
END_DATA_BLOCK

// folder: 20. Robot Services/Tooling & Parking

DATA_BLOCK "ToolChangePepa"   // DB11
{ S7_Optimized_Access := 'TRUE' }
VERSION : 0.1
// stored: InstanceOfName ToolChange
"ToolChange"
BEGIN
END_DATA_BLOCK

DATA_BLOCK "MpsDockingStation_DB"   // DB22
{ S7_Optimized_Access := 'TRUE' }
VERSION : 0.1
// stored: InstanceOfName MpsDockingStation
"MpsDockingStation"
BEGIN
END_DATA_BLOCK

DATA_BLOCK "ToolChangePole_DB"   // DB23
{ S7_Optimized_Access := 'TRUE' }
VERSION : 0.1
// stored: InstanceOfName ToolChange
"ToolChange"
BEGIN
END_DATA_BLOCK

DATA_BLOCK "ToolInRobot_DB"   // DB32
{ S7_Optimized_Access := 'TRUE' }
VERSION : 0.1
// stored: InstanceOfName ToolInRobot
"ToolInRobot"
BEGIN
END_DATA_BLOCK

DATA_BLOCK "ToolChangeGocator_DB"   // DB39
{ S7_Optimized_Access := 'TRUE' }